(* Logix 5000 project; controller PLC_MCC1300_75F1 vendor 1 type 14 code 166 rev 32.11; software revision 32.04; part 72 of 83 *)
(* tags used below, declared in another part *)
   Const_Empty_Data : UDT_Convoy_SL;
   GP_InvertCapxLite : GP_InvertCapxLite;
   GP_OB_InitializeMain : GP_OB_Initialize;
   GP_RampSpace : GP_RampSpace;
   GP_ScadaPlate : GP_ScadaPlate;
   Gp_SpaceConvUtilities_V1 : GP_SpaceConvUtilities_V1;
   M350Popup : MAC_Popup_ZC;
   M350Popup_SL_DATA : UDT_Convoy_SL;
   M351 : MAC_Conveyor;
   M351_ALM : MAC_Conveyor_ALM;
   M351_Data : UDT_Convoy_SL;
   M351_HMR : MAC_Conveyor_HMR;
   M351_HMW : MAC_Conveyor_HMW;
   M351_M1_DR : AXIS_CIP_DRIVE;
   M351_SpaceConv_Utilities : SpaceConv_Utilities;
   M352 : MAC_Conveyor;
   M352_Data : UDT_Convoy_SL;
   M352_SpaceConv_Utilities : SpaceConv_Utilities;
   O : INT[128];
   TMP_d : DINT;
   TMP_dConveyorNumberForZoneCleaning : DINT;
   TMP_dDecelerationPositionEndConveyor : DINT;
   TMP_dOffsetLoadUnload_cmm : DINT;
   TMP_SendToCullet : BOOL;
   TMP_xConveyorInvolvedInCleaning : BOOL;
   TMP_xConveyorOfStartCleaning : BOOL;
   TMP_xEnableLoadUnload : BOOL;
   TMP_xEnableZoneCleaning : BOOL;
   xAlwaysOFF : BOOL;
   xAlwaysON : BOOL;
   Z900 : MAC_Zone;
   Z900_HMI_rgtPlateScada_Internal : HMI_LiteData[5,2,7];
   Z900_HMR : MAC_Zone_HMR;
   Z900_HMW : MAC_Zone_HMW;
(* MainProgram, continued *)

ROUTINE M351_Alarm   (* ladder *)
   // Reset Alarm
   0: XIC(Z900.tmON_ResetAlarm.DN)FLL(0,M351_ALM,1);
   1: XIC(Z900.ST_xEnableControlError)XIC(xAlwaysOFF)XIO(M351.INPUT_xProtectionMotor_M2)OTL(M351_ALM.rgxStoppingFault_M[0].10);
   2: XIC(Z900.ST_xEnableControlError)XIC(M351.INPUT_xDriveError_M2)OTL(M351_ALM.rgxStoppingFault_M[0].11);
   3: XIC(Z900.ST_xEnableControlError)XIO(M351.INPUT_xDriveError_M2)[XIC(M351.OUTPUT_xRun_M2) ,XIC(M351.OUTPUT_xReverse_M2) ,XIC(M351.OUTPUT_xPositioning_M2) ]XIO(M351.INPUT_xDriveFeedback_M2)[XIO(M351.tmON_FeedbackTimeOut_M2.DN) TON(M351.tmON_FeedbackTimeOut_M2,?,?) ,XIC(M351.tmON_FeedbackTimeOut_M2.DN) OTL(M351_ALM.rgxStoppingFault_M[0].12) ];
   4: XIC(Z900.ST_xEnableControlError)XIC(xAlwaysOFF)XIO(M351.INPUT_xLocalSafetySwitch_M2)OTL(M351_ALM.rgxStoppingFault_M[0].13);
   5: XIC(Z900.ST_xEnableControlError)XIO(M351.INPUT_xMotorThermalProbe_M2)OTL(M351_ALM.rgxStoppingFault_M[0].14);
   6: XIC(Z900.ST_xEnableControlError)XIC(xAlwaysOFF)XIO(M351.INPUT_xBrakingResistor_M2)OTL(M351_ALM.rgxStoppingFault_M[0].15);
   7: XIC(Z900.ST_xEnableControlError)XIC(xAlwaysOFF)[XIC(M351.INPUT_xDriveInhibit_M2) ,XIC(M351.OUTPUT_xDriveEnable_M2) XIO(M351.INPUT_xDriveReady_M2) ]OTL(M351_ALM.rgxStoppingFault_M[0].16);
   8: XIC(M351.ST_xEnableControlError)XIC(xAlwaysOFF)XIC(M351.PH_x.7)NEQ(M351_SpaceConv_Utilities.CONST_dSyncMode,0)[XIO(M351.ST_xPlateSynchronized) OTL(M351_ALM.rgxWarning[0].0) ,XIC(M351.ST_xPlateSynchronized) OTU(M351_ALM.rgxWarning[0].0) ];
   9: XIC(M351.ST_xEnableControlError)XIC(xAlwaysOFF)XIC(M351.PH_x.7)XIC(M351_Data.tFlag.tConveyor.xReqStop)OTL(M351_ALM.rgxWarning[0].1);
   // #####_CUMULATIVE ALARM_#####
   10: NOP();
   11: [NEQ(M351_ALM.rgxStoppingFault[0],0) ,NEQ(M351_ALM.rgxStoppingFault_M[0],0) ,NEQ(M351_ALM.rgxStoppingFault_M[1],0) ]OTE(M351.ST_xStopMachineFault);
   12: [NEQ(M351_ALM.rgxFault[0],0) ,NEQ(M351_ALM.rgxFault_M[0],0) ,NEQ(M351_ALM.rgxFault_M[1],0) ]OTE(M351.ST_xStopNextCycleFault);
END_ROUTINE

ROUTINE M351_Logic   (* ladder *)
   // #####_COSTANTS_#####
   0: [MOV(3230,TMP_dConveyorNumberForZoneCleaning) MOV(50000,TMP_dOffsetLoadUnload_cmm) MOV(500,M351_SpaceConv_Utilities.CONST_dPresetFeedbackTime_ms) OTU(TMP_xEnableLoadUnload) OTL(TMP_xEnableZoneCleaning) MOV(450000,M351_SpaceConv_Utilities.CONST_dConveyorLength_cmm) MOV(354800,M351_SpaceConv_Utilities.CONST_dConveyorWidth_cmm) SUB(M351_SpaceConv_Utilities.CONST_dConveyorLength_cmm,M351.AUX_dAccSpace_cmm,M351.AUX_dPresetStopLoad_cmm) ADD(M351_SpaceConv_Utilities.CONST_dConveyorLength_cmm,M351.AUX_dDecSpace_cmm,M351.AUX_dPresetStopUnload_cmm) MOV(1.4,M351_SpaceConv_Utilities.CONST_rAcceleration_ms2) MOV(1.4,M351_SpaceConv_Utilities.CONST_rDeceleration_ms2) ,[MOV(1,M351_SpaceConv_Utilities.CONST_dSyncMode) ,MOV(0,M351_SpaceConv_Utilities.CONST_dSyncroPhPosition_cmm) ,MOV(100000,M351_SpaceConv_Utilities.CONST_dSyncroPhWindow_cmm) ] ];
   // #####_MATCH_#####
   1: NOP();
   // Conveyor Cleaning
   2: XIC(TMP_xEnableZoneCleaning)XIC(Z900.ST_xCleaningAccepted)GRT(Z900_HMW.dCleaningSelection,0)[EQU(Z900_HMW.dCleaningSelection,TMP_dConveyorNumberForZoneCleaning) OTE(TMP_xConveyorOfStartCleaning) ,GEQ(Z900_HMW.dCleaningSelection,TMP_dConveyorNumberForZoneCleaning) OTE(TMP_xConveyorInvolvedInCleaning) ];
   // Enable control error
   3: XIC(Z900.ST_xEnableControlError)OTE(M351.ST_xEnableControlError);
   // Mode 7 - Offsett for load/unload Simultaney
   4: XIC(M351.PH_x.8)MOV(M351.AUX_dPresetStopLoad_cmm,M351_SpaceConv_Utilities.ST_dStopLoadForseen_cmm)MOV(TMP_dOffsetLoadUnload_cmm,M351_SpaceConv_Utilities.CONF_MD7_dOffset_cmm)GP_SpaceConvUtilities_V1(Gp_SpaceConvUtilities_V1,M351_SpaceConv_Utilities,M351_SpaceConv_Utilities,M352_SpaceConv_Utilities,7);
   // #####_ALARMS_#####
   5: NOP();
   // Call Alarm Routine
   6: JSR(M351_Alarm,0);
   // #####_HMI_LOGICS_#####
   7: NOP();
   // Condition ok for Cleaning
   8: [XIO(TMP_xEnableZoneCleaning) ,XIC(TMP_xEnableZoneCleaning) [XIC(M351.ST_xOutputEnable) ,XIO(xAlwaysOFF) ] [XIO(TMP_xConveyorOfStartCleaning) ,XIC(M351.PH_x.0) ,XIO(M351.PH_x.8) ] ]OTE(M351.ST_xCleaningConditionOK);
   // Cleaning Accepted
   9: [XIC(M351_HMW.xStopLocalCleaningRequest) OTU(M351_HMW.xStopLocalCleaningRequest) OTU(M351_HMW.xLocalCleaningRequest) ,XIC(M351_HMW.xLocalCleaningRequest) [XIC(M351.ST_xCleaningConditionOK) ,XIC(M351.ST_xCleaningAccepted) ] OTE(M351.ST_xCleaningAccepted) ];
   // Manual Mode Enabled
   10: XIO(M351_SpaceConv_Utilities.ST_xFeedbackRotation)[XIC(M351_HMW.xEnableDisableManualCommand) XIC(M350Popup.INPUT_xPopupHigh) XIC(M351.ST_xConditionOKStopCycle) OTL(M351.ST_xManualMode) ,[XIO(M351_HMW.xEnableDisableManualCommand) ,XIO(M350Popup.INPUT_xPopupHigh) ] OTU(M351.ST_xManualMode) ];
   // Virtual door enabled
   11: XIC(M351_HMW.xEnableDisableVirtualDoor)OTE(M351.ST_xVirtualDoorEnabled);
   // Clear manual command
   12: XIO(M351.ST_xManualMode)MOV(0,M351_HMW.rgxMan);
   // #####_STATUSES_#####
   13: NOP();
   // Machine in Alarm
   14: [XIC(M351.ST_xStopMachineFault) ,XIC(M351.ST_xStopNextCycleFault) ]OTE(M351.ST_xMachineAlarm);
   // Condition ok for stop Cycle
   15: [XIO(M351.ST_xPhasesInProgress) ,XIC(M351.PH_x.8) XIO(M351.OUTPUT_xRun_M2) XIO(M351_SpaceConv_Utilities.ST_xFeedbackRotation) ,XIC(M351.ST_xMachineAlarm) ,XIO(Z900.ST_xCycleON) ]OTE(M351.ST_xConditionOKStopCycle);
   // Cycle load unload simultaneous
   16: XIC(TMP_xEnableLoadUnload)XIO(M351.ST_xDisableLoadUnloadOnStop)XIO(M351.ST_xIdPlatePresence)OTE(M351.ST_xCycleLoadUnload);
   // Speed Management
   17: [XIO(M351_SpaceConv_Utilities.O_xRampInProgress) XIO(M351.ST_xManualMode) MOV(Z900_HMR.dLineSpeed_mm_min,M351.AUX_dReqSpeed_mm_min) ,[XIC(M351.PH_x.0) ,XIC(M351.PH_x.24) ] MOV(M352.AUX_dReqSpeed_mm_min,M351.AUX_dReqSpeed_mm_min) ,XIC(M351.ST_xManualMode) MOV(Z900_HMW.dManualSpeed_mm_min,M351.AUX_dReqSpeed_mm_min) ,NEQ(M351.AUX_dReqSpeed_mm_min,M351_SpaceConv_Utilities.ST_dRealSpeed_mm_min) OTE(M351.OS_xChangeSpeed) ];
   // Ramp Management
   18: GP_RampSpace(GP_RampSpace,M351_SpaceConv_Utilities.CONST_rAcceleration_ms2,M351_SpaceConv_Utilities.CONST_rDeceleration_ms2,M351_SpaceConv_Utilities.ST_dRealSpeed_mm_min,M351.AUX_dAccSpace_cmm,M351.AUX_dDecSpace_cmm);
   // Space Convoy utilities MOD 1 for Calculate Head/Tail
   19: XIC(xAlwaysON)[[XIC(M351.OUTPUT_xRun_M2) ,XIC(M351.OUTPUT_xReverse_M2) ] XIO(M351.ST_xManualMode) OTE(M351_SpaceConv_Utilities.CONF_MD1_xRun) ,XIC(M351.OUTPUT_xReverse_M2) XIC(xAlwaysOFF) XIO(M351.ST_xManualMode) OTE(M351_SpaceConv_Utilities.CONF_MD1_xReverse) ,[XIC(M351.INPUT_xDriveFeedback_M2) ,XIC(M351_SpaceConv_Utilities.CONF_MD1_xRun) GRT(M351_SpaceConv_Utilities.O_dCountFeedbackTime_ms,0) ] OTE(M351_SpaceConv_Utilities.ST_xFeedbackRotation) ,XIC(M351.ST_xIdPlatePresence) OTE(M351_SpaceConv_Utilities.CONF_MD1_xHeadTracking) ,XIC(M351.ST_xPlatePresence) OTE(M351_SpaceConv_Utilities.CONF_MD1_xTailTracking) ,MOV(GP_OB_InitializeMain.OUT_dExecutionTime_ms,M351_SpaceConv_Utilities.CONF_MD1_dScan_ms) GP_SpaceConvUtilities_V1(Gp_SpaceConvUtilities_V1,M351_SpaceConv_Utilities,M351_SpaceConv_Utilities,M352_SpaceConv_Utilities,1) ];
   // Output Enable
   20: XIC(Z900.ST_xCycleON)XIO(M351.ST_xManualMode)XIO(M351.ST_xStopMachineFault)[XIO(M351.ST_xPlatePassageUpstream_FW) XIO(M351.ST_xPlatePassageUpstream_BKW) ,XIC(M351.ST_xPlatePassageUpstream_FW) XIC(M352.ST_xOutputEnable) ,XIC(M351.ST_xPlatePassageUpstream_BKW) XIC(xAlwaysOFF) ]XIC(M351.INPUT_xHighPositionPopup_1)OTE(M351.ST_xOutputEnable);
   // #####_WORKING_FLAGS_#####
   21: NOP();
   // #####_LOGICS_#####
   22: NOP();
   // Phase of load (from sample)
   23: XIC(M352.OS_xUnload_FW)[OTL(M351.PH_x.0) ,OTU(M351_SpaceConv_Utilities.O_xPlateSynchronized) ,OTU(M351.ST_xDisableLoadUnloadOnStop) ,OTE(M351.OS_xLoad_FW) ,COP(M352_Data,M351_Data,1) FLL(0,M352_Data,1) ,GP_SpaceConvUtilities_V1(Gp_SpaceConvUtilities_V1,M351_SpaceConv_Utilities,M352_SpaceConv_Utilities,M351_SpaceConv_Utilities,5) ];
   // End load Phase (from sample)
   24: XIC(M351.PH_x.0)[GRT(M351_SpaceConv_Utilities.O_dHeadPosition_cmm,M351.AUX_dPresetStopLoad_cmm) ,CPT(TMP_d,M351_Data.dLength_cmm / 2 + M351_SpaceConv_Utilities.CONST_dConveyorWidth_cmm / 2) GRT(M351_SpaceConv_Utilities.O_dHeadPosition_cmm,TMP_d) ][OTE(M351.PH_x.7) ,OTU(M351.PH_x.0) ,OTL(M351.ST_xPlatePresence) ];
   // New data received from MainLine
   25: XIC(M351.ST_xAux4)XIC(M350Popup.AUX_tSearchPlateData.xPlateHooked)XIC(M350Popup.PH_xEndRise)[GP_InvertCapxLite(GP_InvertCapxLite,0,0,0,M350Popup_SL_DATA,M351_Data,Const_Empty_Data,M351_SpaceConv_Utilities.CONST_dConveyorWidth_cmm,M351_SpaceConv_Utilities.CONST_dConveyorLength_cmm,M351_SpaceConv_Utilities.CONF_MD2_MD3_dPrstPos_cmm,M350Popup.AUX_dPosition_cmm,200000) ,GP_SpaceConvUtilities_V1(Gp_SpaceConvUtilities_V1,M351_SpaceConv_Utilities,M351_SpaceConv_Utilities,M352_SpaceConv_Utilities,2) ,OTL(M351.ST_xPlatePresence) ];
   // Calculation Space for Wait Stop Next Conveyor
   26: CPT(TMP_dDecelerationPositionEndConveyor,M351_SpaceConv_Utilities.CONST_dConveyorLength_cmm - M351.AUX_dAccSpace_cmm + 1000);
   // Wait stop next Machine
   27: XIO(M351.PH_x.8)GEQ(M351_SpaceConv_Utilities.O_dHeadPosition_cmm,TMP_dDecelerationPositionEndConveyor)OTE(M351.ST_xWaitStopNextMachine);
   // Set Wait Machine Stop
   28: [XIC(M351.PH_x.7) [XIO(M352.ST_xInitialConditionOK) ,XIC(M351.ST_xWaitStopNextMachine) [XIC(M352_SpaceConv_Utilities.O_xRampInProgress) ,XIO(M352_SpaceConv_Utilities.ST_xFeedbackRotation) ] ] ,XIC(M351.PH_x.0) NEQ(Z900_HMR.dLineSpeed_mm_min,M351.AUX_dReqSpeed_mm_min) ]OTL(M351.ST_xWaitMachineStop);
   // Reset Wait Machine Stop
   29: XIO(M351_SpaceConv_Utilities.ST_xFeedbackRotation)[XIO(M351_SpaceConv_Utilities.ST_xFeedbackRotation) ,XIO(M351.ST_xWaitStopNextMachine) ]EQU(Z900_HMR.dLineSpeed_mm_min,M351.AUX_dReqSpeed_mm_min)OTU(M351.ST_xWaitMachineStop);
   // Phase of unload (to sample)
   30: XIC(Z900.ST_xConditionOkPhaseAdvancement)XIC(M351.ST_xPlatePresence)XIC(M351.ST_xIdPlatePresence)XIC(M351.ST_xOutputEnable)XIC(M352.ST_xInitialConditionOK)XIO(M351.ST_xWaitMachineStop)XIO(M351.PH_x.8)[OTE(M351.ST_xWaitReadyToMove) ,[XIC(M351.ST_xAxleReadyToMoveDelayed) ,XIC(xAlwaysON) ] [OTE(M351.OS_xUnload_FW) ,OTL(M351.PH_x.8) ,MOV(M351_Data.dLength_cmm,M351_SpaceConv_Utilities.CONF_MD4_MD6_dLength_cmm) GP_SpaceConvUtilities_V1(Gp_SpaceConvUtilities_V1,M351_SpaceConv_Utilities,M351_SpaceConv_Utilities,M352_SpaceConv_Utilities,6) ] ];
   // Phase of end unload (to sample)
   31: XIC(M351.PH_x.8)[GEQ(M351_SpaceConv_Utilities.O_dTailPosition_cmm,M351.AUX_dPresetStopUnload_cmm) ,[XIO(M351_SpaceConv_Utilities.ST_xFeedbackRotation) ,XIO(xAlwaysOFF) ] GEQ(M351_SpaceConv_Utilities.O_dTailPosition_cmm,M351_SpaceConv_Utilities.CONST_dConveyorLength_cmm) ][OTE(M351.PH_x.15) ,OTU(M351.PH_x.8) ,OTU(M351.ST_xPlatePresence) ];
   // Phase in progress
   32: NEQ(M351.PH_x,0)OTE(M351.ST_xPhasesInProgress);
   // #####_CLEANING_#####
   33: NOP();
   // Cleaning Reset
   34: XIC(M351.ST_xCleaningAccepted)[XIC(Z900.ST_xCleaningAccepted) ,XIO(TMP_xConveyorOfStartCleaning) ][XIC(M351.ST_xIdPlatePresence) OTL(TMP_SendToCullet) FLL(0,M351_Data,1) ,MOV(0,M351.PH_x) OTU(M351.ST_xPlatePresence) ];
   // Initial condition OK (sample)
   35: XIC(Z900.ST_xConditionOkPhaseAdvancement)XIC(M351.ST_xOutputEnable)XIO(M351_HMW.xEnableDisableManualCommand)XIO(M351.ST_xReqCleaning)XIO(M351.ST_xCleaningAccepted)XIO(M351.ST_xStopNextCycleFault)XIO(M351.ST_xVirtualDoorEnabled)XIO(M352.ST_xVirtualDoorEnabled)XIO(M351.PH_x.0)[XIO(M351.ST_xPhasesInProgress) XIO(M351.ST_xPlatePresence) ,XIC(M351.ST_xCycleLoadUnload) XIC(M351.PH_x.8) [XIC(M351.OUTPUT_xRun_M2) ,XIC(M351.OUTPUT_xRun_M3) ] GRT(M351_SpaceConv_Utilities.O_dTailPosition_cmm,M351_SpaceConv_Utilities.O_dPresetLoadUnload_cmm) XIO(M351.ST_xIdPlatePresence) ]OTE(M351.ST_xInitialConditionOK);
   // #####_HMI_STATUSES_#####
   36: NOP();
   // Manual Mode Enable {x|x|x|x|O}
   37: XIC(M351.ST_xManualMode)OTE(M351_HMR.xManualCommandEnabled);
   // Command forward M2
   38: XIC(M351.ST_xManualMode)XIC(M351_HMW.rgxMan.2)XIC(M351.OUTPUT_xRun_M2)OTE(M351_HMR.rgxMan.2);
   // Command backward M2
   39: XIC(M351.ST_xManualMode)XIC(M351_HMW.rgxMan.3)XIC(M351.OUTPUT_xReverse_M2)OTE(M351_HMR.rgxMan.3);
   // Cleaning Enabled {x|x|x|x|O}
   40: XIC(M351.ST_xCleaningAccepted)[XIC(Z900.ST_xCleaningAccepted) ,XIO(TMP_xEnableZoneCleaning) ]OTE(M351_HMR.xCleaningEnabled);
   // Virtual door Enabled {x|x|x|x|O}
   41: XIC(M351.ST_xVirtualDoorEnabled)OTE(M351_HMR.xVirtualDoorEnabled);
   // Id plate presence
   42: XIC(M351.ST_xIdPlatePresence)OTE(M351_HMR.xIdPlatePresence);
   // Machine state M2
   43: XIC(xAlwaysON)[MOV(1,M351_HMR.dState2) ,XIC(M351.OUTPUT_xRun_M2) MOV(3,M351_HMR.dState2) ,XIC(M351.OUTPUT_xReverse_M2) MOV(4,M351_HMR.dState2) ,XIC(M351.ST_xMachineAlarm) MOV(7,M351_HMR.dState2) ];
   44: XIC(M351_SpaceConv_Utilities.O_xPlateSynchronized)OTE(M351.ST_xPlateSynchronized);
   // State Sensor
   45: XIC(xAlwaysON)[MOV(1,M351_HMR.dStateSensor1) ,XIC(M351_ALM.rgxWarning[0].0) MOV(7,M351_HMR.dStateSensor1) ];
   // Motor error code
   46: MOV(M351_M1_DR.AxisFault,M351_HMR.dErrorCode2);
   47: XIC(M351.ST_xIdPlatePresence)GP_ScadaPlate(GP_ScadaPlate,M351_Data,0,M351_SpaceConv_Utilities.O_dHeadPosition_cmm,M351_SpaceConv_Utilities.CONST_dConveyorWidth_cmm,M351_SpaceConv_Utilities.CONST_dConveyorLength_cmm,M351_SpaceConv_Utilities.ST_xLastModLoadBkw,M351_SpaceConv_Utilities.ST_xLastModUnloadBkw,1,1,Z900_HMI_rgtPlateScada_Internal);
END_ROUTINE
